   4238: 'Carrier 66 Encoder Internal Error', class No Acknowledgement, trigger "DB302_HMI_Faults_Carrier66_Faults_0" bit 13
   4239: 'Carrier 66 Encoder Comm Fault', class No Acknowledgement, trigger "DB302_HMI_Faults_Carrier66_Faults_0" bit 14
   4240: 'Carrier 66 HMI Comm Fault', class No Acknowledgement, trigger "DB302_HMI_Faults_Carrier66_Faults_0" bit 15
   4241: 'Carrier 66 Crash Detection Fault', class No Acknowledgement, trigger "DB302_HMI_Faults_Carrier66_Faults_1" bit 0
   4242: 'Carrier 66 Carrier Number Invalid', class No Acknowledgement, trigger "DB302_HMI_Faults_Carrier66_Faults_1" bit 1
   4243: 'Carrier 66 Drive: PROFINET configuration error', class No Acknowledgement, trigger "DB302_HMI_Faults_Carrier66_Faults_1" bit 2
   4244: 'Carrier 66 Drive: Error internal communications', class No Acknowledgement, trigger "DB302_HMI_Faults_Carrier66_Faults_1" bit 3
   4245: 'Carrier 66 Drive: Motor overtemperature', class No Acknowledgement, trigger "DB302_HMI_Faults_Carrier66_Faults_1" bit 4
   4246: 'Carrier 66 Drive: Motor overcurrent', class No Acknowledgement, trigger "DB302_HMI_Faults_Carrier66_Faults_1" bit 5
   4247: 'Carrier 66 Drive: Infeed or power unit not ready', class No Acknowledgement, trigger "DB302_HMI_Faults_Carrier66_Faults_1" bit 6
   4248: 'Carrier 66 Drive: Short-circuit/ground fault detected', class No Acknowledgement, trigger "DB302_HMI_Faults_Carrier66_Faults_1" bit 7
   4249: 'Carrier 66 Drive: PROFINET Setpoint timeout', class No Acknowledgement, trigger "DB302_HMI_Faults_Carrier66_Faults_1" bit 8
   4250: 'Carrier 66 Power unit: Overcurrent', class No Acknowledgement, trigger "DB302_HMI_Faults_Carrier66_Faults_1" bit 9
   4251: 'Carrier 66 Power unit: DC link voltage overvoltage', class No Acknowledgement, trigger "DB302_HMI_Faults_Carrier66_Faults_1" bit 10
   4252: 'Carrier 66 Power unit: DC link voltage undervoltage', class No Acknowledgement, trigger "DB302_HMI_Faults_Carrier66_Faults_1" bit 11
   4253: 'Carrier 66 Power unit: Line phase failure in main circuit', class No Acknowledgement, trigger "DB302_HMI_Faults_Carrier66_Faults_1" bit 12
   4254: 'Carrier 66 Power unit: Phase failure motor cable', class No Acknowledgement, trigger "DB302_HMI_Faults_Carrier66_Faults_1" bit 13
   4255: 'Carrier 66 Power unit: Ground fault', class No Acknowledgement, trigger "DB302_HMI_Faults_Carrier66_Faults_1" bit 14
   4256: 'Spare_Fault_4256', class No Acknowledgement, trigger "DB302_HMI_Faults_Carrier66_Faults_1" bit 15
   4257: 'Carrier 66 Motion Off Fault', class No Acknowledgement, trigger "DB302_HMI_Faults_Carrier66_Faults_2" bit 0
   4258: 'Carrier 66 Motion On Fault', class No Acknowledgement, trigger "DB302_HMI_Faults_Carrier66_Faults_2" bit 1
   4259: 'Carrier 66 Spacing Fault', class No Acknowledgement, trigger "DB302_HMI_Faults_Carrier66_Faults_2" bit 2
   4260: 'Carrier 66 Duplicate Carrier Number Fault', class No Acknowledgement, trigger "DB302_HMI_Faults_Carrier66_Faults_2" bit 3
   4261: 'Spare_Fault_4261', class No Acknowledgement, trigger "DB302_HMI_Faults_Carrier66_Faults_2" bit 4
   4262: 'Spare_Fault_4262', class No Acknowledgement, trigger "DB302_HMI_Faults_Carrier66_Faults_2" bit 5
   4263: 'Spare_Fault_4263', class No Acknowledgement, trigger "DB302_HMI_Faults_Carrier66_Faults_2" bit 6
   4264: 'Spare_Fault_4264', class No Acknowledgement, trigger "DB302_HMI_Faults_Carrier66_Faults_2" bit 7
   4265: 'Spare_Fault_4265', class No Acknowledgement, trigger "DB302_HMI_Faults_Carrier66_Faults_2" bit 8
   4266: 'Spare_Fault_4266', class No Acknowledgement, trigger "DB302_HMI_Faults_Carrier66_Faults_2" bit 9
   4267: 'Spare_Fault_4267', class No Acknowledgement, trigger "DB302_HMI_Faults_Carrier66_Faults_2" bit 10
   4268: 'Spare_Fault_4268', class No Acknowledgement, trigger "DB302_HMI_Faults_Carrier66_Faults_2" bit 11
   4269: 'Spare_Fault_4269', class No Acknowledgement, trigger "DB302_HMI_Faults_Carrier66_Faults_2" bit 12
   4270: 'Spare_Fault_4270', class No Acknowledgement, trigger "DB302_HMI_Faults_Carrier66_Faults_2" bit 13
   4271: 'Spare_Fault_4271', class No Acknowledgement, trigger "DB302_HMI_Faults_Carrier66_Faults_2" bit 14
   4272: 'Spare_Fault_4272', class No Acknowledgement, trigger "DB302_HMI_Faults_Carrier66_Faults_2" bit 15
   4273: 'Spare_Fault_4273', class No Acknowledgement, trigger "DB302_HMI_Faults_Carrier66_Faults_3" bit 0
   4274: 'Spare_Fault_4274', class No Acknowledgement, trigger "DB302_HMI_Faults_Carrier66_Faults_3" bit 1
   4275: 'Spare_Fault_4275', class No Acknowledgement, trigger "DB302_HMI_Faults_Carrier66_Faults_3" bit 2
   4276: 'Spare_Fault_4276', class No Acknowledgement, trigger "DB302_HMI_Faults_Carrier66_Faults_3" bit 3
   4277: 'Spare_Fault_4277', class No Acknowledgement, trigger "DB302_HMI_Faults_Carrier66_Faults_3" bit 4
   4278: 'Spare_Fault_4278', class No Acknowledgement, trigger "DB302_HMI_Faults_Carrier66_Faults_3" bit 5
   4279: 'Spare_Fault_4279', class No Acknowledgement, trigger "DB302_HMI_Faults_Carrier66_Faults_3" bit 6
   4280: 'Spare_Fault_4280', class No Acknowledgement, trigger "DB302_HMI_Faults_Carrier66_Faults_3" bit 7
   4281: 'Spare_Fault_4281', class No Acknowledgement, trigger "DB302_HMI_Faults_Carrier66_Faults_3" bit 8
   4282: 'Spare_Fault_4282', class No Acknowledgement, trigger "DB302_HMI_Faults_Carrier66_Faults_3" bit 9
   4283: 'Spare_Fault_4283', class No Acknowledgement, trigger "DB302_HMI_Faults_Carrier66_Faults_3" bit 10
   4284: 'Spare_Fault_4284', class No Acknowledgement, trigger "DB302_HMI_Faults_Carrier66_Faults_3" bit 11
   4285: 'Spare_Fault_4285', class No Acknowledgement, trigger "DB302_HMI_Faults_Carrier66_Faults_3" bit 12
   4286: 'Spare_Fault_4286', class No Acknowledgement, trigger "DB302_HMI_Faults_Carrier66_Faults_3" bit 13
   4287: 'Spare_Fault_4287', class No Acknowledgement, trigger "DB302_HMI_Faults_Carrier66_Faults_3" bit 14
   4288: 'Spare_Fault_4288', class No Acknowledgement, trigger "DB302_HMI_Faults_Carrier66_Faults_3" bit 15
   4289: 'Carrier 67 Disconnect Open Power Fault DI11.0', class No Acknowledgement, trigger "DB302_HMI_Faults_Carrier67_Faults_0" bit 0
   4290: 'Carrier 67 Drive Profinet Comm Fault', class No Acknowledgement, trigger "DB302_HMI_Faults_Carrier67_Faults_0" bit 1
   4291: 'Carrier 67 Production Stop Not Reset', class No Acknowledgement, trigger "DB302_HMI_Faults_Carrier67_Faults_0" bit 2
   4292: 'Carrier 67 CB02122 Tripped', class No Acknowledgement, trigger "DB302_HMI_Faults_Carrier67_Faults_0" bit 3
   4293: 'Carrier 67 CB02123 Tripped', class No Acknowledgement, trigger "DB302_HMI_Faults_Carrier67_Faults_0" bit 4
   4294: 'Carrier 67 AUX1 CB Tripped', class No Acknowledgement, trigger "DB302_HMI_Faults_Carrier67_Faults_0" bit 5
   4295: 'Carrier 67 AUX2 CB Tripped', class No Acknowledgement, trigger "DB302_HMI_Faults_Carrier67_Faults_0" bit 6
   4296: 'Carrier 67 PLC Not Communicating', class No Acknowledgement, trigger "DB302_HMI_Faults_Carrier67_Faults_0" bit 7
   4297: 'Carrier 67 Safe Input Card Fault', class No Acknowledgement, trigger "DB302_HMI_Faults_Carrier67_Faults_0" bit 8
   4298: 'Carrier 67 Safe Output Card Fault', class No Acknowledgement, trigger "DB302_HMI_Faults_Carrier67_Faults_0" bit 9
   4299: 'Carrier 67 Standard Input Card Fault', class No Acknowledgement, trigger "DB302_HMI_Faults_Carrier67_Faults_0" bit 10
   4300: 'Carrier 67 Standard Output Card Fault', class No Acknowledgement, trigger "DB302_HMI_Faults_Carrier67_Faults_0" bit 11
   4301: 'Carrier 67 Encoder Position Fault', class No Acknowledgement, trigger "DB302_HMI_Faults_Carrier67_Faults_0" bit 12
   4302: 'Carrier 67 Encoder Internal Error', class No Acknowledgement, trigger "DB302_HMI_Faults_Carrier67_Faults_0" bit 13
   4303: 'Carrier 67 Encoder Comm Fault', class No Acknowledgement, trigger "DB302_HMI_Faults_Carrier67_Faults_0" bit 14
   4304: 'Carrier 67 HMI Comm Fault', class No Acknowledgement, trigger "DB302_HMI_Faults_Carrier67_Faults_0" bit 15
   4305: 'Carrier 67 Crash Detection Fault', class No Acknowledgement, trigger "DB302_HMI_Faults_Carrier67_Faults_1" bit 0
   4306: 'Carrier 67 Carrier Number Invalid', class No Acknowledgement, trigger "DB302_HMI_Faults_Carrier67_Faults_1" bit 1
   4307: 'Carrier 67 Drive: PROFINET configuration error', class No Acknowledgement, trigger "DB302_HMI_Faults_Carrier67_Faults_1" bit 2
   4308: 'Carrier 67 Drive: Error internal communications', class No Acknowledgement, trigger "DB302_HMI_Faults_Carrier67_Faults_1" bit 3
   4309: 'Carrier 67 Drive: Motor overtemperature', class No Acknowledgement, trigger "DB302_HMI_Faults_Carrier67_Faults_1" bit 4
   4310: 'Carrier 67 Drive: Motor overcurrent', class No Acknowledgement, trigger "DB302_HMI_Faults_Carrier67_Faults_1" bit 5
   4311: 'Carrier 67 Drive: Infeed or power unit not ready', class No Acknowledgement, trigger "DB302_HMI_Faults_Carrier67_Faults_1" bit 6
   4312: 'Carrier 67 Drive: Short-circuit/ground fault detected', class No Acknowledgement, trigger "DB302_HMI_Faults_Carrier67_Faults_1" bit 7
   4313: 'Carrier 67 Drive: PROFINET Setpoint timeout', class No Acknowledgement, trigger "DB302_HMI_Faults_Carrier67_Faults_1" bit 8
   4314: 'Carrier 67 Power unit: Overcurrent', class No Acknowledgement, trigger "DB302_HMI_Faults_Carrier67_Faults_1" bit 9
   4315: 'Carrier 67 Power unit: DC link voltage overvoltage', class No Acknowledgement, trigger "DB302_HMI_Faults_Carrier67_Faults_1" bit 10
   4316: 'Carrier 67 Power unit: DC link voltage undervoltage', class No Acknowledgement, trigger "DB302_HMI_Faults_Carrier67_Faults_1" bit 11
   4317: 'Carrier 67 Power unit: Line phase failure in main circuit', class No Acknowledgement, trigger "DB302_HMI_Faults_Carrier67_Faults_1" bit 12
   4318: 'Carrier 67 Power unit: Phase failure motor cable', class No Acknowledgement, trigger "DB302_HMI_Faults_Carrier67_Faults_1" bit 13
   4319: 'Carrier 67 Power unit: Ground fault', class No Acknowledgement, trigger "DB302_HMI_Faults_Carrier67_Faults_1" bit 14
   4320: 'Spare_Fault_4320', class No Acknowledgement, trigger "DB302_HMI_Faults_Carrier67_Faults_1" bit 15
   4321: 'Carrier 67 Motion Off Fault', class No Acknowledgement, trigger "DB302_HMI_Faults_Carrier67_Faults_2" bit 0
   4322: 'Carrier 67 Motion On Fault', class No Acknowledgement, trigger "DB302_HMI_Faults_Carrier67_Faults_2" bit 1
   4323: 'Carrier 67 Spacing Fault', class No Acknowledgement, trigger "DB302_HMI_Faults_Carrier67_Faults_2" bit 2
   4324: 'Carrier 67 Duplicate Carrier Number Fault', class No Acknowledgement, trigger "DB302_HMI_Faults_Carrier67_Faults_2" bit 3
   4325: 'Spare_Fault_4325', class No Acknowledgement, trigger "DB302_HMI_Faults_Carrier67_Faults_2" bit 4
   4326: 'Spare_Fault_4326', class No Acknowledgement, trigger "DB302_HMI_Faults_Carrier67_Faults_2" bit 5
   4327: 'Spare_Fault_4327', class No Acknowledgement, trigger "DB302_HMI_Faults_Carrier67_Faults_2" bit 6
   4328: 'Spare_Fault_4328', class No Acknowledgement, trigger "DB302_HMI_Faults_Carrier67_Faults_2" bit 7
   4329: 'Spare_Fault_4329', class No Acknowledgement, trigger "DB302_HMI_Faults_Carrier67_Faults_2" bit 8
   4330: 'Spare_Fault_4330', class No Acknowledgement, trigger "DB302_HMI_Faults_Carrier67_Faults_2" bit 9
   4331: 'Spare_Fault_4331', class No Acknowledgement, trigger "DB302_HMI_Faults_Carrier67_Faults_2" bit 10
   4332: 'Spare_Fault_4332', class No Acknowledgement, trigger "DB302_HMI_Faults_Carrier67_Faults_2" bit 11
   4333: 'Spare_Fault_4333', class No Acknowledgement, trigger "DB302_HMI_Faults_Carrier67_Faults_2" bit 12
   4334: 'Spare_Fault_4334', class No Acknowledgement, trigger "DB302_HMI_Faults_Carrier67_Faults_2" bit 13
   4335: 'Spare_Fault_4335', class No Acknowledgement, trigger "DB302_HMI_Faults_Carrier67_Faults_2" bit 14
   4336: 'Spare_Fault_4336', class No Acknowledgement, trigger "DB302_HMI_Faults_Carrier67_Faults_2" bit 15
   4337: 'Spare_Fault_4337', class No Acknowledgement, trigger "DB302_HMI_Faults_Carrier67_Faults_3" bit 0
   4338: 'Spare_Fault_4338', class No Acknowledgement, trigger "DB302_HMI_Faults_Carrier67_Faults_3" bit 1
   4339: 'Spare_Fault_4339', class No Acknowledgement, trigger "DB302_HMI_Faults_Carrier67_Faults_3" bit 2
   4340: 'Spare_Fault_4340', class No Acknowledgement, trigger "DB302_HMI_Faults_Carrier67_Faults_3" bit 3
   4341: 'Spare_Fault_4341', class No Acknowledgement, trigger "DB302_HMI_Faults_Carrier67_Faults_3" bit 4
   4342: 'Spare_Fault_4342', class No Acknowledgement, trigger "DB302_HMI_Faults_Carrier67_Faults_3" bit 5
   4343: 'Spare_Fault_4343', class No Acknowledgement, trigger "DB302_HMI_Faults_Carrier67_Faults_3" bit 6
   4344: 'Spare_Fault_4344', class No Acknowledgement, trigger "DB302_HMI_Faults_Carrier67_Faults_3" bit 7
   4345: 'Spare_Fault_4345', class No Acknowledgement, trigger "DB302_HMI_Faults_Carrier67_Faults_3" bit 8
   4346: 'Spare_Fault_4346', class No Acknowledgement, trigger "DB302_HMI_Faults_Carrier67_Faults_3" bit 9
   4347: 'Spare_Fault_4347', class No Acknowledgement, trigger "DB302_HMI_Faults_Carrier67_Faults_3" bit 10
   4348: 'Spare_Fault_4348', class No Acknowledgement, trigger "DB302_HMI_Faults_Carrier67_Faults_3" bit 11
   4349: 'Spare_Fault_4349', class No Acknowledgement, trigger "DB302_HMI_Faults_Carrier67_Faults_3" bit 12
   4350: 'Spare_Fault_4350', class No Acknowledgement, trigger "DB302_HMI_Faults_Carrier67_Faults_3" bit 13
   4351: 'Spare_Fault_4351', class No Acknowledgement, trigger "DB302_HMI_Faults_Carrier67_Faults_3" bit 14
   4352: 'Spare_Fault_4352', class No Acknowledgement, trigger "DB302_HMI_Faults_Carrier67_Faults_3" bit 15
   4353: 'Carrier 68 Disconnect Open Power Fault DI11.0', class No Acknowledgement, trigger "DB302_HMI_Faults_Carrier68_Faults_0" bit 0
   4354: 'Carrier 68 Drive Profinet Comm Fault', class No Acknowledgement, trigger "DB302_HMI_Faults_Carrier68_Faults_0" bit 1
   4355: 'Carrier 68 Production Stop Not Reset', class No Acknowledgement, trigger "DB302_HMI_Faults_Carrier68_Faults_0" bit 2
   4356: 'Carrier 68 CB02122 Tripped', class No Acknowledgement, trigger "DB302_HMI_Faults_Carrier68_Faults_0" bit 3
   4357: 'Carrier 68 CB02123 Tripped', class No Acknowledgement, trigger "DB302_HMI_Faults_Carrier68_Faults_0" bit 4
   4358: 'Carrier 68 AUX1 CB Tripped', class No Acknowledgement, trigger "DB302_HMI_Faults_Carrier68_Faults_0" bit 5
   4359: 'Carrier 68 AUX2 CB Tripped', class No Acknowledgement, trigger "DB302_HMI_Faults_Carrier68_Faults_0" bit 6
   4360: 'Carrier 68 PLC Not Communicating', class No Acknowledgement, trigger "DB302_HMI_Faults_Carrier68_Faults_0" bit 7
   4361: 'Carrier 68 Safe Input Card Fault', class No Acknowledgement, trigger "DB302_HMI_Faults_Carrier68_Faults_0" bit 8
   4362: 'Carrier 68 Safe Output Card Fault', class No Acknowledgement, trigger "DB302_HMI_Faults_Carrier68_Faults_0" bit 9
   4363: 'Carrier 68 Standard Input Card Fault', class No Acknowledgement, trigger "DB302_HMI_Faults_Carrier68_Faults_0" bit 10
   4364: 'Carrier 68 Standard Output Card Fault', class No Acknowledgement, trigger "DB302_HMI_Faults_Carrier68_Faults_0" bit 11
   4365: 'Carrier 68 Encoder Position Fault', class No Acknowledgement, trigger "DB302_HMI_Faults_Carrier68_Faults_0" bit 12
   4366: 'Carrier 68 Encoder Internal Error', class No Acknowledgement, trigger "DB302_HMI_Faults_Carrier68_Faults_0" bit 13
   4367: 'Carrier 68 Encoder Comm Fault', class No Acknowledgement, trigger "DB302_HMI_Faults_Carrier68_Faults_0" bit 14
   4368: 'Carrier 68 HMI Comm Fault', class No Acknowledgement, trigger "DB302_HMI_Faults_Carrier68_Faults_0" bit 15
   4369: 'Carrier 68 Crash Detection Fault', class No Acknowledgement, trigger "DB302_HMI_Faults_Carrier68_Faults_1" bit 0
   4370: 'Carrier 68 Carrier Number Invalid', class No Acknowledgement, trigger "DB302_HMI_Faults_Carrier68_Faults_1" bit 1
   4371: 'Carrier 68 Drive: PROFINET configuration error', class No Acknowledgement, trigger "DB302_HMI_Faults_Carrier68_Faults_1" bit 2
   4372: 'Carrier 68 Drive: Error internal communications', class No Acknowledgement, trigger "DB302_HMI_Faults_Carrier68_Faults_1" bit 3
   4373: 'Carrier 68 Drive: Motor overtemperature', class No Acknowledgement, trigger "DB302_HMI_Faults_Carrier68_Faults_1" bit 4
   4374: 'Carrier 68 Drive: Motor overcurrent', class No Acknowledgement, trigger "DB302_HMI_Faults_Carrier68_Faults_1" bit 5
   4375: 'Carrier 68 Drive: Infeed or power unit not ready', class No Acknowledgement, trigger "DB302_HMI_Faults_Carrier68_Faults_1" bit 6
   4376: 'Carrier 68 Drive: Short-circuit/ground fault detected', class No Acknowledgement, trigger "DB302_HMI_Faults_Carrier68_Faults_1" bit 7
   4377: 'Carrier 68 Drive: PROFINET Setpoint timeout', class No Acknowledgement, trigger "DB302_HMI_Faults_Carrier68_Faults_1" bit 8
   4378: 'Carrier 68 Power unit: Overcurrent', class No Acknowledgement, trigger "DB302_HMI_Faults_Carrier68_Faults_1" bit 9
   4379: 'Carrier 68 Power unit: DC link voltage overvoltage', class No Acknowledgement, trigger "DB302_HMI_Faults_Carrier68_Faults_1" bit 10
   4380: 'Carrier 68 Power unit: DC link voltage undervoltage', class No Acknowledgement, trigger "DB302_HMI_Faults_Carrier68_Faults_1" bit 11
   4381: 'Carrier 68 Power unit: Line phase failure in main circuit', class No Acknowledgement, trigger "DB302_HMI_Faults_Carrier68_Faults_1" bit 12
   4382: 'Carrier 68 Power unit: Phase failure motor cable', class No Acknowledgement, trigger "DB302_HMI_Faults_Carrier68_Faults_1" bit 13
   4383: 'Carrier 68 Power unit: Ground fault', class No Acknowledgement, trigger "DB302_HMI_Faults_Carrier68_Faults_1" bit 14
   4384: 'Spare_Fault_4384', class No Acknowledgement, trigger "DB302_HMI_Faults_Carrier68_Faults_1" bit 15
   4385: 'Carrier 68 Motion Off Fault', class No Acknowledgement, trigger "DB302_HMI_Faults_Carrier68_Faults_2" bit 0
   4386: 'Carrier 68 Motion On Fault', class No Acknowledgement, trigger "DB302_HMI_Faults_Carrier68_Faults_2" bit 1
   4387: 'Carrier 68 Spacing Fault', class No Acknowledgement, trigger "DB302_HMI_Faults_Carrier68_Faults_2" bit 2
   4388: 'Carrier 68 Duplicate Carrier Number Fault', class No Acknowledgement, trigger "DB302_HMI_Faults_Carrier68_Faults_2" bit 3
   4389: 'Spare_Fault_4389', class No Acknowledgement, trigger "DB302_HMI_Faults_Carrier68_Faults_2" bit 4
   4390: 'Spare_Fault_4390', class No Acknowledgement, trigger "DB302_HMI_Faults_Carrier68_Faults_2" bit 5
   4391: 'Spare_Fault_4391', class No Acknowledgement, trigger "DB302_HMI_Faults_Carrier68_Faults_2" bit 6
   4392: 'Spare_Fault_4392', class No Acknowledgement, trigger "DB302_HMI_Faults_Carrier68_Faults_2" bit 7
   4393: 'Spare_Fault_4393', class No Acknowledgement, trigger "DB302_HMI_Faults_Carrier68_Faults_2" bit 8
   4394: 'Spare_Fault_4394', class No Acknowledgement, trigger "DB302_HMI_Faults_Carrier68_Faults_2" bit 9
   4395: 'Spare_Fault_4395', class No Acknowledgement, trigger "DB302_HMI_Faults_Carrier68_Faults_2" bit 10
   4396: 'Spare_Fault_4396', class No Acknowledgement, trigger "DB302_HMI_Faults_Carrier68_Faults_2" bit 11
   4397: 'Spare_Fault_4397', class No Acknowledgement, trigger "DB302_HMI_Faults_Carrier68_Faults_2" bit 12
   4398: 'Spare_Fault_4398', class No Acknowledgement, trigger "DB302_HMI_Faults_Carrier68_Faults_2" bit 13
   4399: 'Spare_Fault_4399', class No Acknowledgement, trigger "DB302_HMI_Faults_Carrier68_Faults_2" bit 14
   4400: 'Spare_Fault_4400', class No Acknowledgement, trigger "DB302_HMI_Faults_Carrier68_Faults_2" bit 15
   4401: 'Spare_Fault_4401', class No Acknowledgement, trigger "DB302_HMI_Faults_Carrier68_Faults_3" bit 0
   4402: 'Spare_Fault_4402', class No Acknowledgement, trigger "DB302_HMI_Faults_Carrier68_Faults_3" bit 1
   4403: 'Spare_Fault_4403', class No Acknowledgement, trigger "DB302_HMI_Faults_Carrier68_Faults_3" bit 2
   4404: 'Spare_Fault_4404', class No Acknowledgement, trigger "DB302_HMI_Faults_Carrier68_Faults_3" bit 3
   4405: 'Spare_Fault_4405', class No Acknowledgement, trigger "DB302_HMI_Faults_Carrier68_Faults_3" bit 4
   4406: 'Spare_Fault_4406', class No Acknowledgement, trigger "DB302_HMI_Faults_Carrier68_Faults_3" bit 5
   4407: 'Spare_Fault_4407', class No Acknowledgement, trigger "DB302_HMI_Faults_Carrier68_Faults_3" bit 6
   4408: 'Spare_Fault_4408', class No Acknowledgement, trigger "DB302_HMI_Faults_Carrier68_Faults_3" bit 7
   4409: 'Spare_Fault_4409', class No Acknowledgement, trigger "DB302_HMI_Faults_Carrier68_Faults_3" bit 8
   4410: 'Spare_Fault_4410', class No Acknowledgement, trigger "DB302_HMI_Faults_Carrier68_Faults_3" bit 9
   4411: 'Spare_Fault_4411', class No Acknowledgement, trigger "DB302_HMI_Faults_Carrier68_Faults_3" bit 10
   4412: 'Spare_Fault_4412', class No Acknowledgement, trigger "DB302_HMI_Faults_Carrier68_Faults_3" bit 11
   4413: 'Spare_Fault_4413', class No Acknowledgement, trigger "DB302_HMI_Faults_Carrier68_Faults_3" bit 12
   4414: 'Spare_Fault_4414', class No Acknowledgement, trigger "DB302_HMI_Faults_Carrier68_Faults_3" bit 13
   4415: 'Spare_Fault_4415', class No Acknowledgement, trigger "DB302_HMI_Faults_Carrier68_Faults_3" bit 14
   4416: 'Spare_Fault_4416', class No Acknowledgement, trigger "DB302_HMI_Faults_Carrier68_Faults_3" bit 15
   4417: 'Carrier 69 Disconnect Open Power Fault DI11.0', class No Acknowledgement, trigger "DB302_HMI_Faults_Carrier69_Faults_0" bit 0
   4418: 'Carrier 69 Drive Profinet Comm Fault', class No Acknowledgement, trigger "DB302_HMI_Faults_Carrier69_Faults_0" bit 1
   4419: 'Carrier 69 Production Stop Not Reset', class No Acknowledgement, trigger "DB302_HMI_Faults_Carrier69_Faults_0" bit 2
   4420: 'Carrier 69 CB02122 Tripped', class No Acknowledgement, trigger "DB302_HMI_Faults_Carrier69_Faults_0" bit 3
   4421: 'Carrier 69 CB02123 Tripped', class No Acknowledgement, trigger "DB302_HMI_Faults_Carrier69_Faults_0" bit 4
   4422: 'Carrier 69 AUX1 CB Tripped', class No Acknowledgement, trigger "DB302_HMI_Faults_Carrier69_Faults_0" bit 5
   4423: 'Carrier 69 AUX2 CB Tripped', class No Acknowledgement, trigger "DB302_HMI_Faults_Carrier69_Faults_0" bit 6
   4424: 'Carrier 69 PLC Not Communicating', class No Acknowledgement, trigger "DB302_HMI_Faults_Carrier69_Faults_0" bit 7
   4425: 'Carrier 69 Safe Input Card Fault', class No Acknowledgement, trigger "DB302_HMI_Faults_Carrier69_Faults_0" bit 8
   4426: 'Carrier 69 Safe Output Card Fault', class No Acknowledgement, trigger "DB302_HMI_Faults_Carrier69_Faults_0" bit 9
   4427: 'Carrier 69 Standard Input Card Fault', class No Acknowledgement, trigger "DB302_HMI_Faults_Carrier69_Faults_0" bit 10
   4428: 'Carrier 69 Standard Output Card Fault', class No Acknowledgement, trigger "DB302_HMI_Faults_Carrier69_Faults_0" bit 11
   4429: 'Carrier 69 Encoder Position Fault', class No Acknowledgement, trigger "DB302_HMI_Faults_Carrier69_Faults_0" bit 12
   4430: 'Carrier 69 Encoder Internal Error', class No Acknowledgement, trigger "DB302_HMI_Faults_Carrier69_Faults_0" bit 13
   4431: 'Carrier 69 Encoder Comm Fault', class No Acknowledgement, trigger "DB302_HMI_Faults_Carrier69_Faults_0" bit 14
   4432: 'Carrier 69 HMI Comm Fault', class No Acknowledgement, trigger "DB302_HMI_Faults_Carrier69_Faults_0" bit 15
   4433: 'Carrier 69 Crash Detection Fault', class No Acknowledgement, trigger "DB302_HMI_Faults_Carrier69_Faults_1" bit 0
   4434: 'Carrier 69 Carrier Number Invalid', class No Acknowledgement, trigger "DB302_HMI_Faults_Carrier69_Faults_1" bit 1
   4435: 'Carrier 69 Drive: PROFINET configuration error', class No Acknowledgement, trigger "DB302_HMI_Faults_Carrier69_Faults_1" bit 2
   4436: 'Carrier 69 Drive: Error internal communications', class No Acknowledgement, trigger "DB302_HMI_Faults_Carrier69_Faults_1" bit 3
   4437: 'Carrier 69 Drive: Motor overtemperature', class No Acknowledgement, trigger "DB302_HMI_Faults_Carrier69_Faults_1" bit 4
   4438: 'Carrier 69 Drive: Motor overcurrent', class No Acknowledgement, trigger "DB302_HMI_Faults_Carrier69_Faults_1" bit 5
   4439: 'Carrier 69 Drive: Infeed or power unit not ready', class No Acknowledgement, trigger "DB302_HMI_Faults_Carrier69_Faults_1" bit 6
   4440: 'Carrier 69 Drive: Short-circuit/ground fault detected', class No Acknowledgement, trigger "DB302_HMI_Faults_Carrier69_Faults_1" bit 7
   4441: 'Carrier 69 Drive: PROFINET Setpoint timeout', class No Acknowledgement, trigger "DB302_HMI_Faults_Carrier69_Faults_1" bit 8
   4442: 'Carrier 69 Power unit: Overcurrent', class No Acknowledgement, trigger "DB302_HMI_Faults_Carrier69_Faults_1" bit 9
   4443: 'Carrier 69 Power unit: DC link voltage overvoltage', class No Acknowledgement, trigger "DB302_HMI_Faults_Carrier69_Faults_1" bit 10
   4444: 'Carrier 69 Power unit: DC link voltage undervoltage', class No Acknowledgement, trigger "DB302_HMI_Faults_Carrier69_Faults_1" bit 11
   4445: 'Carrier 69 Power unit: Line phase failure in main circuit', class No Acknowledgement, trigger "DB302_HMI_Faults_Carrier69_Faults_1" bit 12
   4446: 'Carrier 69 Power unit: Phase failure motor cable', class No Acknowledgement, trigger "DB302_HMI_Faults_Carrier69_Faults_1" bit 13
   4447: 'Carrier 69 Power unit: Ground fault', class No Acknowledgement, trigger "DB302_HMI_Faults_Carrier69_Faults_1" bit 14
   4448: 'Spare_Fault_4448', class No Acknowledgement, trigger "DB302_HMI_Faults_Carrier69_Faults_1" bit 15
   4449: 'Carrier 69 Motion Off Fault', class No Acknowledgement, trigger "DB302_HMI_Faults_Carrier69_Faults_2" bit 0
   4450: 'Carrier 69 Motion On Fault', class No Acknowledgement, trigger "DB302_HMI_Faults_Carrier69_Faults_2" bit 1
   4451: 'Carrier 69 Spacing Fault', class No Acknowledgement, trigger "DB302_HMI_Faults_Carrier69_Faults_2" bit 2
   4452: 'Carrier 69 Duplicate Carrier Number Fault', class No Acknowledgement, trigger "DB302_HMI_Faults_Carrier69_Faults_2" bit 3
   4453: 'Spare_Fault_4453', class No Acknowledgement, trigger "DB302_HMI_Faults_Carrier69_Faults_2" bit 4
   4454: 'Spare_Fault_4454', class No Acknowledgement, trigger "DB302_HMI_Faults_Carrier69_Faults_2" bit 5
   4455: 'Spare_Fault_4455', class No Acknowledgement, trigger "DB302_HMI_Faults_Carrier69_Faults_2" bit 6
   4456: 'Spare_Fault_4456', class No Acknowledgement, trigger "DB302_HMI_Faults_Carrier69_Faults_2" bit 7
   4457: 'Spare_Fault_4457', class No Acknowledgement, trigger "DB302_HMI_Faults_Carrier69_Faults_2" bit 8
   4458: 'Spare_Fault_4458', class No Acknowledgement, trigger "DB302_HMI_Faults_Carrier69_Faults_2" bit 9
   4459: 'Spare_Fault_4459', class No Acknowledgement, trigger "DB302_HMI_Faults_Carrier69_Faults_2" bit 10
   4460: 'Spare_Fault_4460', class No Acknowledgement, trigger "DB302_HMI_Faults_Carrier69_Faults_2" bit 11
   4461: 'Spare_Fault_4461', class No Acknowledgement, trigger "DB302_HMI_Faults_Carrier69_Faults_2" bit 12
   4462: 'Spare_Fault_4462', class No Acknowledgement, trigger "DB302_HMI_Faults_Carrier69_Faults_2" bit 13
   4463: 'Spare_Fault_4463', class No Acknowledgement, trigger "DB302_HMI_Faults_Carrier69_Faults_2" bit 14
   4464: 'Spare_Fault_4464', class No Acknowledgement, trigger "DB302_HMI_Faults_Carrier69_Faults_2" bit 15
   4465: 'Spare_Fault_4465', class No Acknowledgement, trigger "DB302_HMI_Faults_Carrier69_Faults_3" bit 0
   4466: 'Spare_Fault_4466', class No Acknowledgement, trigger "DB302_HMI_Faults_Carrier69_Faults_3" bit 1
   4467: 'Spare_Fault_4467', class No Acknowledgement, trigger "DB302_HMI_Faults_Carrier69_Faults_3" bit 2
   4468: 'Spare_Fault_4468', class No Acknowledgement, trigger "DB302_HMI_Faults_Carrier69_Faults_3" bit 3
   4469: 'Spare_Fault_4469', class No Acknowledgement, trigger "DB302_HMI_Faults_Carrier69_Faults_3" bit 4
   4470: 'Spare_Fault_4470', class No Acknowledgement, trigger "DB302_HMI_Faults_Carrier69_Faults_3" bit 5
   4471: 'Spare_Fault_4471', class No Acknowledgement, trigger "DB302_HMI_Faults_Carrier69_Faults_3" bit 6
   4472: 'Spare_Fault_4472', class No Acknowledgement, trigger "DB302_HMI_Faults_Carrier69_Faults_3" bit 7
   4473: 'Spare_Fault_4473', class No Acknowledgement, trigger "DB302_HMI_Faults_Carrier69_Faults_3" bit 8
   4474: 'Spare_Fault_4474', class No Acknowledgement, trigger "DB302_HMI_Faults_Carrier69_Faults_3" bit 9
   4475: 'Spare_Fault_4475', class No Acknowledgement, trigger "DB302_HMI_Faults_Carrier69_Faults_3" bit 10
   4476: 'Spare_Fault_4476', class No Acknowledgement, trigger "DB302_HMI_Faults_Carrier69_Faults_3" bit 11
   4477: 'Spare_Fault_4477', class No Acknowledgement, trigger "DB302_HMI_Faults_Carrier69_Faults_3" bit 12
   4478: 'Spare_Fault_4478', class No Acknowledgement, trigger "DB302_HMI_Faults_Carrier69_Faults_3" bit 13
   4479: 'Spare_Fault_4479', class No Acknowledgement, trigger "DB302_HMI_Faults_Carrier69_Faults_3" bit 14
   4480: 'Spare_Fault_4480', class No Acknowledgement, trigger "DB302_HMI_Faults_Carrier69_Faults_3" bit 15
   4481: 'Carrier 70 Disconnect Open Power Fault DI11.0', class No Acknowledgement, trigger "DB302_HMI_Faults_Carrier70_Faults_0" bit 0
   4482: 'Carrier 70 Drive Profinet Comm Fault', class No Acknowledgement, trigger "DB302_HMI_Faults_Carrier70_Faults_0" bit 1
   4483: 'Carrier 70 Production Stop Not Reset', class No Acknowledgement, trigger "DB302_HMI_Faults_Carrier70_Faults_0" bit 2
   4484: 'Carrier 70 CB02122 Tripped', class No Acknowledgement, trigger "DB302_HMI_Faults_Carrier70_Faults_0" bit 3
   4485: 'Carrier 70 CB02123 Tripped', class No Acknowledgement, trigger "DB302_HMI_Faults_Carrier70_Faults_0" bit 4
   4486: 'Carrier 70 AUX1 CB Tripped', class No Acknowledgement, trigger "DB302_HMI_Faults_Carrier70_Faults_0" bit 5
   4487: 'Carrier 70 AUX2 CB Tripped', class No Acknowledgement, trigger "DB302_HMI_Faults_Carrier70_Faults_0" bit 6
   4488: 'Carrier 70 PLC Not Communicating', class No Acknowledgement, trigger "DB302_HMI_Faults_Carrier70_Faults_0" bit 7
   4489: 'Carrier 70 Safe Input Card Fault', class No Acknowledgement, trigger "DB302_HMI_Faults_Carrier70_Faults_0" bit 8
   4490: 'Carrier 70 Safe Output Card Fault', class No Acknowledgement, trigger "DB302_HMI_Faults_Carrier70_Faults_0" bit 9
   4491: 'Carrier 70 Standard Input Card Fault', class No Acknowledgement, trigger "DB302_HMI_Faults_Carrier70_Faults_0" bit 10
   4492: 'Carrier 70 Standard Output Card Fault', class No Acknowledgement, trigger "DB302_HMI_Faults_Carrier70_Faults_0" bit 11
   4493: 'Carrier 70 Encoder Position Fault', class No Acknowledgement, trigger "DB302_HMI_Faults_Carrier70_Faults_0" bit 12
   4494: 'Carrier 70 Encoder Internal Error', class No Acknowledgement, trigger "DB302_HMI_Faults_Carrier70_Faults_0" bit 13
   4495: 'Carrier 70 Encoder Comm Fault', class No Acknowledgement, trigger "DB302_HMI_Faults_Carrier70_Faults_0" bit 14
   4496: 'Carrier 70 HMI Comm Fault', class No Acknowledgement, trigger "DB302_HMI_Faults_Carrier70_Faults_0" bit 15
   4497: 'Carrier 70 Crash Detection Fault', class No Acknowledgement, trigger "DB302_HMI_Faults_Carrier70_Faults_1" bit 0
   4498: 'Carrier 70 Carrier Number Invalid', class No Acknowledgement, trigger "DB302_HMI_Faults_Carrier70_Faults_1" bit 1
   4499: 'Carrier 70 Drive: PROFINET configuration error', class No Acknowledgement, trigger "DB302_HMI_Faults_Carrier70_Faults_1" bit 2
   4500: 'Carrier 70 Drive: Error internal communications', class No Acknowledgement, trigger "DB302_HMI_Faults_Carrier70_Faults_1" bit 3
   4501: 'Carrier 70 Drive: Motor overtemperature', class No Acknowledgement, trigger "DB302_HMI_Faults_Carrier70_Faults_1" bit 4
   4502: 'Carrier 70 Drive: Motor overcurrent', class No Acknowledgement, trigger "DB302_HMI_Faults_Carrier70_Faults_1" bit 5
   4503: 'Carrier 70 Drive: Infeed or power unit not ready', class No Acknowledgement, trigger "DB302_HMI_Faults_Carrier70_Faults_1" bit 6
   4504: 'Carrier 70 Drive: Short-circuit/ground fault detected', class No Acknowledgement, trigger "DB302_HMI_Faults_Carrier70_Faults_1" bit 7
   4505: 'Carrier 70 Drive: PROFINET Setpoint timeout', class No Acknowledgement, trigger "DB302_HMI_Faults_Carrier70_Faults_1" bit 8
   4506: 'Carrier 70 Power unit: Overcurrent', class No Acknowledgement, trigger "DB302_HMI_Faults_Carrier70_Faults_1" bit 9
   4507: 'Carrier 70 Power unit: DC link voltage overvoltage', class No Acknowledgement, trigger "DB302_HMI_Faults_Carrier70_Faults_1" bit 10
   4508: 'Carrier 70 Power unit: DC link voltage undervoltage', class No Acknowledgement, trigger "DB302_HMI_Faults_Carrier70_Faults_1" bit 11
   4509: 'Carrier 70 Power unit: Line phase failure in main circuit', class No Acknowledgement, trigger "DB302_HMI_Faults_Carrier70_Faults_1" bit 12
   4510: 'Carrier 70 Power unit: Phase failure motor cable', class No Acknowledgement, trigger "DB302_HMI_Faults_Carrier70_Faults_1" bit 13
   4511: 'Carrier 70 Power unit: Ground fault', class No Acknowledgement, trigger "DB302_HMI_Faults_Carrier70_Faults_1" bit 14
   4512: 'Spare_Fault_4512', class No Acknowledgement, trigger "DB302_HMI_Faults_Carrier70_Faults_1" bit 15
   4513: 'Carrier 70 Motion Off Fault', class No Acknowledgement, trigger "DB302_HMI_Faults_Carrier70_Faults_2" bit 0
   4514: 'Carrier 70 Motion On Fault', class No Acknowledgement, trigger "DB302_HMI_Faults_Carrier70_Faults_2" bit 1
   4515: 'Carrier 70 Spacing Fault', class No Acknowledgement, trigger "DB302_HMI_Faults_Carrier70_Faults_2" bit 2
   4516: 'Carrier 70 Duplicate Carrier Number Fault', class No Acknowledgement, trigger "DB302_HMI_Faults_Carrier70_Faults_2" bit 3
   4517: 'Spare_Fault_4517', class No Acknowledgement, trigger "DB302_HMI_Faults_Carrier70_Faults_2" bit 4
   4518: 'Spare_Fault_4518', class No Acknowledgement, trigger "DB302_HMI_Faults_Carrier70_Faults_2" bit 5
   4519: 'Spare_Fault_4519', class No Acknowledgement, trigger "DB302_HMI_Faults_Carrier70_Faults_2" bit 6
   4520: 'Spare_Fault_4520', class No Acknowledgement, trigger "DB302_HMI_Faults_Carrier70_Faults_2" bit 7
   4521: 'Spare_Fault_4521', class No Acknowledgement, trigger "DB302_HMI_Faults_Carrier70_Faults_2" bit 8
   4522: 'Spare_Fault_4522', class No Acknowledgement, trigger "DB302_HMI_Faults_Carrier70_Faults_2" bit 9
   4523: 'Spare_Fault_4523', class No Acknowledgement, trigger "DB302_HMI_Faults_Carrier70_Faults_2" bit 10
   4524: 'Spare_Fault_4524', class No Acknowledgement, trigger "DB302_HMI_Faults_Carrier70_Faults_2" bit 11
   4525: 'Spare_Fault_4525', class No Acknowledgement, trigger "DB302_HMI_Faults_Carrier70_Faults_2" bit 12
   4526: 'Spare_Fault_4526', class No Acknowledgement, trigger "DB302_HMI_Faults_Carrier70_Faults_2" bit 13
   4527: 'Spare_Fault_4527', class No Acknowledgement, trigger "DB302_HMI_Faults_Carrier70_Faults_2" bit 14
   4528: 'Spare_Fault_4528', class No Acknowledgement, trigger "DB302_HMI_Faults_Carrier70_Faults_2" bit 15
   4529: 'Spare_Fault_4529', class No Acknowledgement, trigger "DB302_HMI_Faults_Carrier70_Faults_3" bit 0
   4530: 'Spare_Fault_4530', class No Acknowledgement, trigger "DB302_HMI_Faults_Carrier70_Faults_3" bit 1
   4531: 'Spare_Fault_4531', class No Acknowledgement, trigger "DB302_HMI_Faults_Carrier70_Faults_3" bit 2
   4532: 'Spare_Fault_4532', class No Acknowledgement, trigger "DB302_HMI_Faults_Carrier70_Faults_3" bit 3
   4533: 'Spare_Fault_4533', class No Acknowledgement, trigger "DB302_HMI_Faults_Carrier70_Faults_3" bit 4
   4534: 'Spare_Fault_4534', class No Acknowledgement, trigger "DB302_HMI_Faults_Carrier70_Faults_3" bit 5
   4535: 'Spare_Fault_4535', class No Acknowledgement, trigger "DB302_HMI_Faults_Carrier70_Faults_3" bit 6
   4536: 'Spare_Fault_4536', class No Acknowledgement, trigger "DB302_HMI_Faults_Carrier70_Faults_3" bit 7
   4537: 'Spare_Fault_4537', class No Acknowledgement, trigger "DB302_HMI_Faults_Carrier70_Faults_3" bit 8
   4538: 'Spare_Fault_4538', class No Acknowledgement, trigger "DB302_HMI_Faults_Carrier70_Faults_3" bit 9
   4539: 'Spare_Fault_4539', class No Acknowledgement, trigger "DB302_HMI_Faults_Carrier70_Faults_3" bit 10
   4540: 'Spare_Fault_4540', class No Acknowledgement, trigger "DB302_HMI_Faults_Carrier70_Faults_3" bit 11
   4541: 'Spare_Fault_4541', class No Acknowledgement, trigger "DB302_HMI_Faults_Carrier70_Faults_3" bit 12
   4542: 'Spare_Fault_4542', class No Acknowledgement, trigger "DB302_HMI_Faults_Carrier70_Faults_3" bit 13
   4543: 'Spare_Fault_4543', class No Acknowledgement, trigger "DB302_HMI_Faults_Carrier70_Faults_3" bit 14
   4544: 'Spare_Fault_4544', class No Acknowledgement, trigger "DB302_HMI_Faults_Carrier70_Faults_3" bit 15
   4545: 'Carrier 71 Disconnect Open Power Fault DI11.0', class No Acknowledgement, trigger "DB302_HMI_Faults_Carrier71_Faults_0" bit 0
   4546: 'Carrier 71 Drive Profinet Comm Fault', class No Acknowledgement, trigger "DB302_HMI_Faults_Carrier71_Faults_0" bit 1
   4547: 'Carrier 71 Production Stop Not Reset', class No Acknowledgement, trigger "DB302_HMI_Faults_Carrier71_Faults_0" bit 2
   4548: 'Carrier 71 CB02122 Tripped', class No Acknowledgement, trigger "DB302_HMI_Faults_Carrier71_Faults_0" bit 3
   4549: 'Carrier 71 CB02123 Tripped', class No Acknowledgement, trigger "DB302_HMI_Faults_Carrier71_Faults_0" bit 4
   4550: 'Carrier 71 AUX1 CB Tripped', class No Acknowledgement, trigger "DB302_HMI_Faults_Carrier71_Faults_0" bit 5
   4551: 'Carrier 71 AUX2 CB Tripped', class No Acknowledgement, trigger "DB302_HMI_Faults_Carrier71_Faults_0" bit 6
   4552: 'Carrier 71 PLC Not Communicating', class No Acknowledgement, trigger "DB302_HMI_Faults_Carrier71_Faults_0" bit 7
   4553: 'Carrier 71 Safe Input Card Fault', class No Acknowledgement, trigger "DB302_HMI_Faults_Carrier71_Faults_0" bit 8
   4554: 'Carrier 71 Safe Output Card Fault', class No Acknowledgement, trigger "DB302_HMI_Faults_Carrier71_Faults_0" bit 9
   4555: 'Carrier 71 Standard Input Card Fault', class No Acknowledgement, trigger "DB302_HMI_Faults_Carrier71_Faults_0" bit 10
   4556: 'Carrier 71 Standard Output Card Fault', class No Acknowledgement, trigger "DB302_HMI_Faults_Carrier71_Faults_0" bit 11
   4557: 'Carrier 71 Encoder Position Fault', class No Acknowledgement, trigger "DB302_HMI_Faults_Carrier71_Faults_0" bit 12
   4558: 'Carrier 71 Encoder Internal Error', class No Acknowledgement, trigger "DB302_HMI_Faults_Carrier71_Faults_0" bit 13
   4559: 'Carrier 71 Encoder Comm Fault', class No Acknowledgement, trigger "DB302_HMI_Faults_Carrier71_Faults_0" bit 14
   4560: 'Carrier 71 HMI Comm Fault', class No Acknowledgement, trigger "DB302_HMI_Faults_Carrier71_Faults_0" bit 15
   4561: 'Carrier 71 Crash Detection Fault', class No Acknowledgement, trigger "DB302_HMI_Faults_Carrier71_Faults_1" bit 0
   4562: 'Carrier 71 Carrier Number Invalid', class No Acknowledgement, trigger "DB302_HMI_Faults_Carrier71_Faults_1" bit 1
   4563: 'Carrier 71 Drive: PROFINET configuration error', class No Acknowledgement, trigger "DB302_HMI_Faults_Carrier71_Faults_1" bit 2
   4564: 'Carrier 71 Drive: Error internal communications', class No Acknowledgement, trigger "DB302_HMI_Faults_Carrier71_Faults_1" bit 3
   4565: 'Carrier 71 Drive: Motor overtemperature', class No Acknowledgement, trigger "DB302_HMI_Faults_Carrier71_Faults_1" bit 4
   4566: 'Carrier 71 Drive: Motor overcurrent', class No Acknowledgement, trigger "DB302_HMI_Faults_Carrier71_Faults_1" bit 5
   4567: 'Carrier 71 Drive: Infeed or power unit not ready', class No Acknowledgement, trigger "DB302_HMI_Faults_Carrier71_Faults_1" bit 6
   4568: 'Carrier 71 Drive: Short-circuit/ground fault detected', class No Acknowledgement, trigger "DB302_HMI_Faults_Carrier71_Faults_1" bit 7
   4569: 'Carrier 71 Drive: PROFINET Setpoint timeout', class No Acknowledgement, trigger "DB302_HMI_Faults_Carrier71_Faults_1" bit 8
   4570: 'Carrier 71 Power unit: Overcurrent', class No Acknowledgement, trigger "DB302_HMI_Faults_Carrier71_Faults_1" bit 9
   4571: 'Carrier 71 Power unit: DC link voltage overvoltage', class No Acknowledgement, trigger "DB302_HMI_Faults_Carrier71_Faults_1" bit 10
   4572: 'Carrier 71 Power unit: DC link voltage undervoltage', class No Acknowledgement, trigger "DB302_HMI_Faults_Carrier71_Faults_1" bit 11
   4573: 'Carrier 71 Power unit: Line phase failure in main circuit', class No Acknowledgement, trigger "DB302_HMI_Faults_Carrier71_Faults_1" bit 12
   4574: 'Carrier 71 Power unit: Phase failure motor cable', class No Acknowledgement, trigger "DB302_HMI_Faults_Carrier71_Faults_1" bit 13
   4575: 'Carrier 71 Power unit: Ground fault', class No Acknowledgement, trigger "DB302_HMI_Faults_Carrier71_Faults_1" bit 14
   4576: 'Spare_Fault_4576', class No Acknowledgement, trigger "DB302_HMI_Faults_Carrier71_Faults_1" bit 15
   4577: 'Carrier 71 Motion Off Fault', class No Acknowledgement, trigger "DB302_HMI_Faults_Carrier71_Faults_2" bit 0
   4578: 'Carrier 71 Motion On Fault', class No Acknowledgement, trigger "DB302_HMI_Faults_Carrier71_Faults_2" bit 1
   4579: 'Carrier 71 Spacing Fault', class No Acknowledgement, trigger "DB302_HMI_Faults_Carrier71_Faults_2" bit 2
   4580: 'Carrier 71 Duplicate Carrier Number Fault', class No Acknowledgement, trigger "DB302_HMI_Faults_Carrier71_Faults_2" bit 3
   4581: 'Spare_Fault_4581', class No Acknowledgement, trigger "DB302_HMI_Faults_Carrier71_Faults_2" bit 4
   4582: 'Spare_Fault_4582', class No Acknowledgement, trigger "DB302_HMI_Faults_Carrier71_Faults_2" bit 5
   4583: 'Spare_Fault_4583', class No Acknowledgement, trigger "DB302_HMI_Faults_Carrier71_Faults_2" bit 6
   4584: 'Spare_Fault_4584', class No Acknowledgement, trigger "DB302_HMI_Faults_Carrier71_Faults_2" bit 7
   4585: 'Spare_Fault_4585', class No Acknowledgement, trigger "DB302_HMI_Faults_Carrier71_Faults_2" bit 8
   4586: 'Spare_Fault_4586', class No Acknowledgement, trigger "DB302_HMI_Faults_Carrier71_Faults_2" bit 9
   4587: 'Spare_Fault_4587', class No Acknowledgement, trigger "DB302_HMI_Faults_Carrier71_Faults_2" bit 10
   4588: 'Spare_Fault_4588', class No Acknowledgement, trigger "DB302_HMI_Faults_Carrier71_Faults_2" bit 11
   4589: 'Spare_Fault_4589', class No Acknowledgement, trigger "DB302_HMI_Faults_Carrier71_Faults_2" bit 12
   4590: 'Spare_Fault_4590', class No Acknowledgement, trigger "DB302_HMI_Faults_Carrier71_Faults_2" bit 13
   4591: 'Spare_Fault_4591', class No Acknowledgement, trigger "DB302_HMI_Faults_Carrier71_Faults_2" bit 14
   4592: 'Spare_Fault_4592', class No Acknowledgement, trigger "DB302_HMI_Faults_Carrier71_Faults_2" bit 15
   4593: 'Spare_Fault_4593', class No Acknowledgement, trigger "DB302_HMI_Faults_Carrier71_Faults_3" bit 0
   4594: 'Spare_Fault_4594', class No Acknowledgement, trigger "DB302_HMI_Faults_Carrier71_Faults_3" bit 1
   4595: 'Spare_Fault_4595', class No Acknowledgement, trigger "DB302_HMI_Faults_Carrier71_Faults_3" bit 2
   4596: 'Spare_Fault_4596', class No Acknowledgement, trigger "DB302_HMI_Faults_Carrier71_Faults_3" bit 3
   4597: 'Spare_Fault_4597', class No Acknowledgement, trigger "DB302_HMI_Faults_Carrier71_Faults_3" bit 4
   4598: 'Spare_Fault_4598', class No Acknowledgement, trigger "DB302_HMI_Faults_Carrier71_Faults_3" bit 5
   4599: 'Spare_Fault_4599', class No Acknowledgement, trigger "DB302_HMI_Faults_Carrier71_Faults_3" bit 6
   4600: 'Spare_Fault_4600', class No Acknowledgement, trigger "DB302_HMI_Faults_Carrier71_Faults_3" bit 7
   4601: 'Spare_Fault_4601', class No Acknowledgement, trigger "DB302_HMI_Faults_Carrier71_Faults_3" bit 8
   4602: 'Spare_Fault_4602', class No Acknowledgement, trigger "DB302_HMI_Faults_Carrier71_Faults_3" bit 9
   4603: 'Spare_Fault_4603', class No Acknowledgement, trigger "DB302_HMI_Faults_Carrier71_Faults_3" bit 10
   4604: 'Spare_Fault_4604', class No Acknowledgement, trigger "DB302_HMI_Faults_Carrier71_Faults_3" bit 11
   4605: 'Spare_Fault_4605', class No Acknowledgement, trigger "DB302_HMI_Faults_Carrier71_Faults_3" bit 12
   4606: 'Spare_Fault_4606', class No Acknowledgement, trigger "DB302_HMI_Faults_Carrier71_Faults_3" bit 13
   4607: 'Spare_Fault_4607', class No Acknowledgement, trigger "DB302_HMI_Faults_Carrier71_Faults_3" bit 14
   4608: 'Spare_Fault_4608', class No Acknowledgement, trigger "DB302_HMI_Faults_Carrier71_Faults_3" bit 15
   4609: 'Carrier 72 Disconnect Open Power Fault DI11.0', class No Acknowledgement, trigger "DB302_HMI_Faults_Carrier72_Faults_0" bit 0
   4610: 'Carrier 72 Drive Profinet Comm Fault', class No Acknowledgement, trigger "DB302_HMI_Faults_Carrier72_Faults_0" bit 1
   4611: 'Carrier 72 Production Stop Not Reset', class No Acknowledgement, trigger "DB302_HMI_Faults_Carrier72_Faults_0" bit 2
   4612: 'Carrier 72 CB02122 Tripped', class No Acknowledgement, trigger "DB302_HMI_Faults_Carrier72_Faults_0" bit 3
   4613: 'Carrier 72 CB02123 Tripped', class No Acknowledgement, trigger "DB302_HMI_Faults_Carrier72_Faults_0" bit 4
   4614: 'Carrier 72 AUX1 CB Tripped', class No Acknowledgement, trigger "DB302_HMI_Faults_Carrier72_Faults_0" bit 5
   4615: 'Carrier 72 AUX2 CB Tripped', class No Acknowledgement, trigger "DB302_HMI_Faults_Carrier72_Faults_0" bit 6
   4616: 'Carrier 72 PLC Not Communicating', class No Acknowledgement, trigger "DB302_HMI_Faults_Carrier72_Faults_0" bit 7
   4617: 'Carrier 72 Safe Input Card Fault', class No Acknowledgement, trigger "DB302_HMI_Faults_Carrier72_Faults_0" bit 8
   4618: 'Carrier 72 Safe Output Card Fault', class No Acknowledgement, trigger "DB302_HMI_Faults_Carrier72_Faults_0" bit 9
   4619: 'Carrier 72 Standard Input Card Fault', class No Acknowledgement, trigger "DB302_HMI_Faults_Carrier72_Faults_0" bit 10
   4620: 'Carrier 72 Standard Output Card Fault', class No Acknowledgement, trigger "DB302_HMI_Faults_Carrier72_Faults_0" bit 11
   4621: 'Carrier 72 Encoder Position Fault', class No Acknowledgement, trigger "DB302_HMI_Faults_Carrier72_Faults_0" bit 12
   4622: 'Carrier 72 Encoder Internal Error', class No Acknowledgement, trigger "DB302_HMI_Faults_Carrier72_Faults_0" bit 13
   4623: 'Carrier 72 Encoder Comm Fault', class No Acknowledgement, trigger "DB302_HMI_Faults_Carrier72_Faults_0" bit 14
   4624: 'Carrier 72 HMI Comm Fault', class No Acknowledgement, trigger "DB302_HMI_Faults_Carrier72_Faults_0" bit 15
   4625: 'Carrier 72 Crash Detection Fault', class No Acknowledgement, trigger "DB302_HMI_Faults_Carrier72_Faults_1" bit 0
   4626: 'Carrier 72 Carrier Number Invalid', class No Acknowledgement, trigger "DB302_HMI_Faults_Carrier72_Faults_1" bit 1
   4627: 'Carrier 72 Drive: PROFINET configuration error', class No Acknowledgement, trigger "DB302_HMI_Faults_Carrier72_Faults_1" bit 2
   4628: 'Carrier 72 Drive: Error internal communications', class No Acknowledgement, trigger "DB302_HMI_Faults_Carrier72_Faults_1" bit 3
   4629: 'Carrier 72 Drive: Motor overtemperature', class No Acknowledgement, trigger "DB302_HMI_Faults_Carrier72_Faults_1" bit 4
   4630: 'Carrier 72 Drive: Motor overcurrent', class No Acknowledgement, trigger "DB302_HMI_Faults_Carrier72_Faults_1" bit 5
   4631: 'Carrier 72 Drive: Infeed or power unit not ready', class No Acknowledgement, trigger "DB302_HMI_Faults_Carrier72_Faults_1" bit 6
   4632: 'Carrier 72 Drive: Short-circuit/ground fault detected', class No Acknowledgement, trigger "DB302_HMI_Faults_Carrier72_Faults_1" bit 7
   4633: 'Carrier 72 Drive: PROFINET Setpoint timeout', class No Acknowledgement, trigger "DB302_HMI_Faults_Carrier72_Faults_1" bit 8
   4634: 'Carrier 72 Power unit: Overcurrent', class No Acknowledgement, trigger "DB302_HMI_Faults_Carrier72_Faults_1" bit 9
   4635: 'Carrier 72 Power unit: DC link voltage overvoltage', class No Acknowledgement, trigger "DB302_HMI_Faults_Carrier72_Faults_1" bit 10
   4636: 'Carrier 72 Power unit: DC link voltage undervoltage', class No Acknowledgement, trigger "DB302_HMI_Faults_Carrier72_Faults_1" bit 11
   4637: 'Carrier 72 Power unit: Line phase failure in main circuit', class No Acknowledgement, trigger "DB302_HMI_Faults_Carrier72_Faults_1" bit 12
   4638: 'Carrier 72 Power unit: Phase failure motor cable', class No Acknowledgement, trigger "DB302_HMI_Faults_Carrier72_Faults_1" bit 13
   4639: 'Carrier 72 Power unit: Ground fault', class No Acknowledgement, trigger "DB302_HMI_Faults_Carrier72_Faults_1" bit 14
   4640: 'Spare_Fault_4640', class No Acknowledgement, trigger "DB302_HMI_Faults_Carrier72_Faults_1" bit 15
   4641: 'Carrier 72 Motion Off Fault', class No Acknowledgement, trigger "DB302_HMI_Faults_Carrier72_Faults_2" bit 0
   4642: 'Carrier 72 Motion On Fault', class No Acknowledgement, trigger "DB302_HMI_Faults_Carrier72_Faults_2" bit 1
   4643: 'Carrier 72 Spacing Fault', class No Acknowledgement, trigger "DB302_HMI_Faults_Carrier72_Faults_2" bit 2
   4644: 'Carrier 72 Duplicate Carrier Number Fault', class No Acknowledgement, trigger "DB302_HMI_Faults_Carrier72_Faults_2" bit 3
   4645: 'Spare_Fault_4645', class No Acknowledgement, trigger "DB302_HMI_Faults_Carrier72_Faults_2" bit 4
   4646: 'Spare_Fault_4646', class No Acknowledgement, trigger "DB302_HMI_Faults_Carrier72_Faults_2" bit 5
   4647: 'Spare_Fault_4647', class No Acknowledgement, trigger "DB302_HMI_Faults_Carrier72_Faults_2" bit 6
   4648: 'Spare_Fault_4648', class No Acknowledgement, trigger "DB302_HMI_Faults_Carrier72_Faults_2" bit 7
   4649: 'Spare_Fault_4649', class No Acknowledgement, trigger "DB302_HMI_Faults_Carrier72_Faults_2" bit 8
   4650: 'Spare_Fault_4650', class No Acknowledgement, trigger "DB302_HMI_Faults_Carrier72_Faults_2" bit 9
   4651: 'Spare_Fault_4651', class No Acknowledgement, trigger "DB302_HMI_Faults_Carrier72_Faults_2" bit 10
   4652: 'Spare_Fault_4652', class No Acknowledgement, trigger "DB302_HMI_Faults_Carrier72_Faults_2" bit 11
   4653: 'Spare_Fault_4653', class No Acknowledgement, trigger "DB302_HMI_Faults_Carrier72_Faults_2" bit 12
   4654: 'Spare_Fault_4654', class No Acknowledgement, trigger "DB302_HMI_Faults_Carrier72_Faults_2" bit 13
   4655: 'Spare_Fault_4655', class No Acknowledgement, trigger "DB302_HMI_Faults_Carrier72_Faults_2" bit 14
   4656: 'Spare_Fault_4656', class No Acknowledgement, trigger "DB302_HMI_Faults_Carrier72_Faults_2" bit 15
   4657: 'Spare_Fault_4657', class No Acknowledgement, trigger "DB302_HMI_Faults_Carrier72_Faults_3" bit 0
   4658: 'Spare_Fault_4658', class No Acknowledgement, trigger "DB302_HMI_Faults_Carrier72_Faults_3" bit 1